(* Logix 5000 project; controller PLC_MCC1300_75F1 vendor 1 type 14 code 166 rev 32.11; software revision 32.04; part 20 of 83 *)
(* tags used below, declared in another part *)
   GP_M311A : GP_Rotator;
   M310B : MAC_Conveyor;
   M311 : MAC_Conveyor;
   M311_ALM : MAC_Conveyor_ALM;
   M311_Data : UDT_Convoy_SL;
   M311_HMR : MAC_Conveyor_HMR;
   M311_HMW : MAC_Conveyor_HMW;
   M311_M1_DR : AXIS_CIP_DRIVE;
   M311_M1_DR_IN_MAJ : MOTION_INSTRUCTION;
   M311_M1_DR_IN_MAR : MOTION_INSTRUCTION;
   M311_M1_DR_IN_MAS : MOTION_INSTRUCTION;
   M311_M1_DR_IN_MRP : MOTION_INSTRUCTION;
   M311_M1_DR_MAFR : MOTION_INSTRUCTION;
   M311_M1_DR_MDR : MOTION_INSTRUCTION;
   M311_M1_DR_MSF : MOTION_INSTRUCTION;
   M311_M1_DR_MSO : MOTION_INSTRUCTION;
   M311_M1_DR_OUT_MAJ : MOTION_INSTRUCTION;
   M311_M1_DR_OUT_MAM : MOTION_INSTRUCTION;
   M311_M1_DR_OUT_MAR : MOTION_INSTRUCTION;
   M311_M1_DR_OUT_MAS : MOTION_INSTRUCTION;
   M311_M1_DR_OUT_MCD : MOTION_INSTRUCTION;
   M311_M1_DR_OUT_MRP : MOTION_INSTRUCTION;
   M311_SpaceConv_Utilities : SpaceConv_Utilities;
   M311A : MAC_Rotator;
   M311A_HMR : MAC_Rotator_HMR;
   M311A_HMW : MAC_Rotator_HMW;
   M311A_M1_DR : AXIS_CIP_DRIVE;
   M311A_M1_DR_IN_MAM : MOTION_INSTRUCTION;
   M311A_M1_DR_IN_MAS : MOTION_INSTRUCTION;
   M311A_M1_DR_MAFR : MOTION_INSTRUCTION;
   M311A_M1_DR_MAH : MOTION_INSTRUCTION;
   M311A_M1_DR_MSF : MOTION_INSTRUCTION;
   M311A_M1_DR_MSO : MOTION_INSTRUCTION;
   M311A_M1_DR_OUT_MAJ : MOTION_INSTRUCTION;
   M311A_M1_DR_OUT_MAM : MOTION_INSTRUCTION;
   M311A_M1_DR_OUT_MAS : MOTION_INSTRUCTION;
   M311A_MAM_IP_TOFF : TIMER;
   M312 : MAC_Conveyor_Single;
   TMP_dDirection : DINT;
   TMP_r : REAL;
   TMP_rAcc : REAL;
   TMP_rDec : REAL;
   TMP_rSpeed : REAL;
   TMP_rTarget : REAL;
   TMP_rTarget_M1 : REAL;
   TMP_xForwardCommadnForCleaningZone : BOOL;
   TMP_xPositioning_M1 : BOOL;
   TMP_xPowerSaving : BOOL;
   TMP_xReverse_M1 : BOOL;
   TMP_xRun_M1 : BOOL;
   xDebugOFF : BOOL;
   Z401 : MAC_Zone;
   Z401_HMW : MAC_Zone_HMW;
(* CommandLogic, continued *)

ROUTINE M311_Output   (* ladder *)
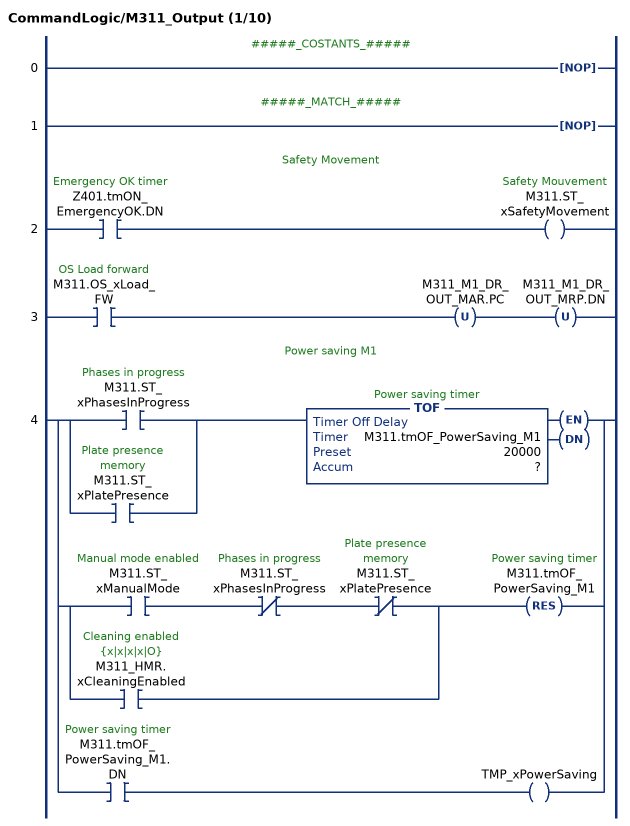
   // #####_COSTANTS_#####
   0: NOP();
   // #####_MATCH_#####
   1: NOP();
   // Safety Movement
   2: XIC(Z401.tmON_EmergencyOK.DN)OTE(M311.ST_xSafetyMovement);
   3: XIC(M311.OS_xLoad_FW)OTU(M311_M1_DR_OUT_MAR.PC)OTU(M311_M1_DR_OUT_MRP.DN);
   // Power saving M1
   4: [[XIC(M311.ST_xPhasesInProgress) ,XIC(M311.ST_xPlatePresence) ] TOF(M311.tmOF_PowerSaving_M1,?,?) ,[XIC(M311.ST_xManualMode) XIO(M311.ST_xPhasesInProgress) XIO(M311.ST_xPlatePresence) ,XIC(M311_HMR.xCleaningEnabled) ] RES(M311.tmOF_PowerSaving_M1) ,XIC(M311.tmOF_PowerSaving_M1.DN) OTE(TMP_xPowerSaving) ];
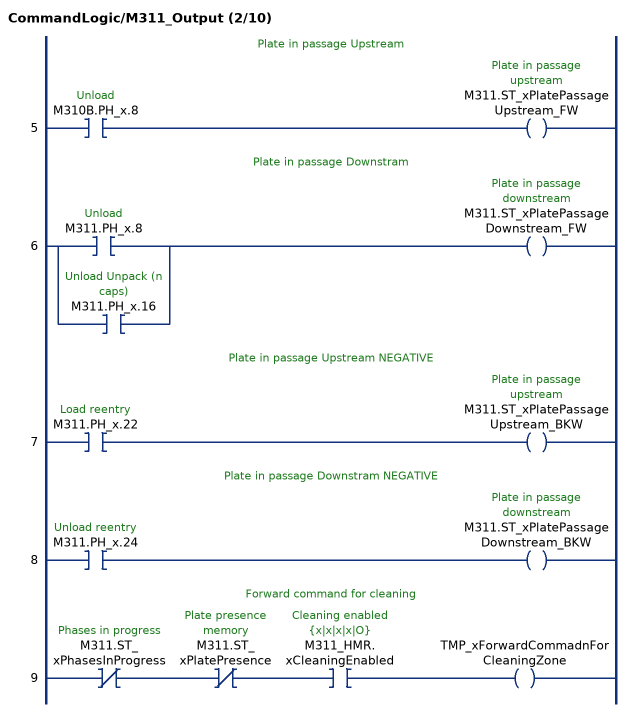
   // Plate in passage Upstream
   5: XIC(M310B.PH_x.8)OTE(M311.ST_xPlatePassageUpstream_FW);
   // Plate in passage Downstram
   6: [XIC(M311.PH_x.8) ,XIC(M311.PH_x.16) ]OTE(M311.ST_xPlatePassageDownstream_FW);
   // Plate in passage Upstream NEGATIVE
   7: XIC(M311.PH_x.22)OTE(M311.ST_xPlatePassageUpstream_BKW);
   // Plate in passage Downstram NEGATIVE
   8: XIC(M311.PH_x.24)OTE(M311.ST_xPlatePassageDownstream_BKW);
   // Forward command for cleaning
   9: XIO(M311.ST_xPhasesInProgress)XIO(M311.ST_xPlatePresence)XIC(M311_HMR.xCleaningEnabled)OTE(TMP_xForwardCommadnForCleaningZone);
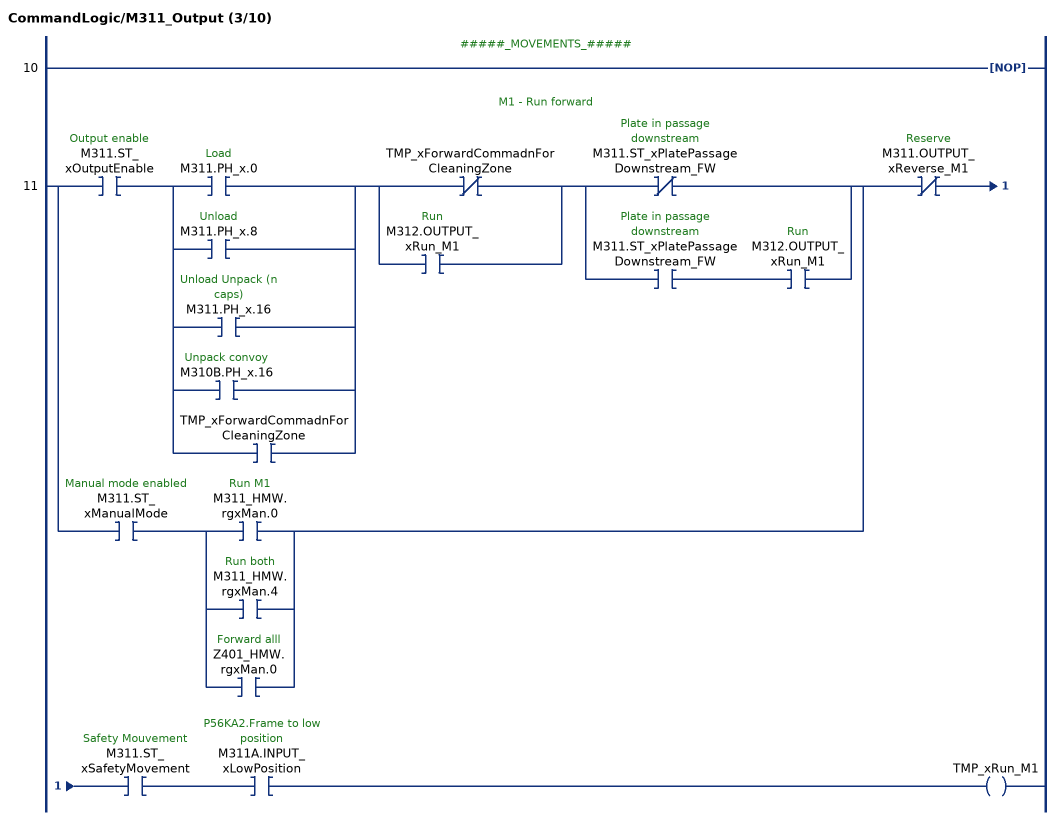
   // #####_MOVEMENTS_#####
   10: NOP();
   // M1 - Run forward
   11: [XIC(M311.ST_xOutputEnable) [XIC(M311.PH_x.0) ,XIC(M311.PH_x.8) ,XIC(M311.PH_x.16) ,XIC(M310B.PH_x.16) ,XIC(TMP_xForwardCommadnForCleaningZone) ] [XIO(TMP_xForwardCommadnForCleaningZone) ,XIC(M312.OUTPUT_xRun_M1) ] [XIO(M311.ST_xPlatePassageDownstream_FW) ,XIC(M311.ST_xPlatePassageDownstream_FW) XIC(M312.OUTPUT_xRun_M1) ] ,XIC(M311.ST_xManualMode) [XIC(M311_HMW.rgxMan.0) ,XIC(M311_HMW.rgxMan.4) ,XIC(Z401_HMW.rgxMan.0) ] ]XIO(M311.OUTPUT_xReverse_M1)XIC(M311.ST_xSafetyMovement)XIC(M311A.INPUT_xLowPosition)OTE(TMP_xRun_M1);
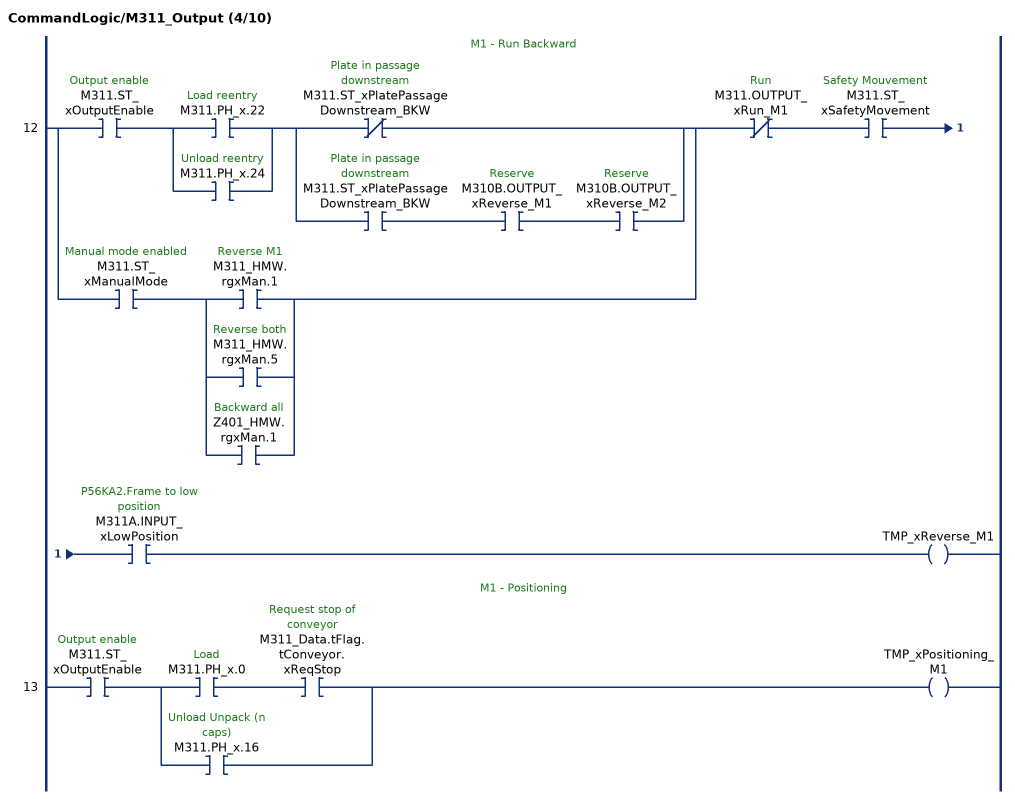
   // M1 - Run Backward
   12: [XIC(M311.ST_xOutputEnable) [XIC(M311.PH_x.22) ,XIC(M311.PH_x.24) ] [XIO(M311.ST_xPlatePassageDownstream_BKW) ,XIC(M311.ST_xPlatePassageDownstream_BKW) XIC(M310B.OUTPUT_xReverse_M1) XIC(M310B.OUTPUT_xReverse_M2) ] ,XIC(M311.ST_xManualMode) [XIC(M311_HMW.rgxMan.1) ,XIC(M311_HMW.rgxMan.5) ,XIC(Z401_HMW.rgxMan.1) ] ]XIO(M311.OUTPUT_xRun_M1)XIC(M311.ST_xSafetyMovement)XIC(M311A.INPUT_xLowPosition)OTE(TMP_xReverse_M1);
   // M1 - Positioning
   13: XIC(M311.ST_xOutputEnable)[XIC(M311.PH_x.0) XIC(M311_Data.tFlag.tConveyor.xReqStop) ,XIC(M311.PH_x.16) ]OTE(TMP_xPositioning_M1);
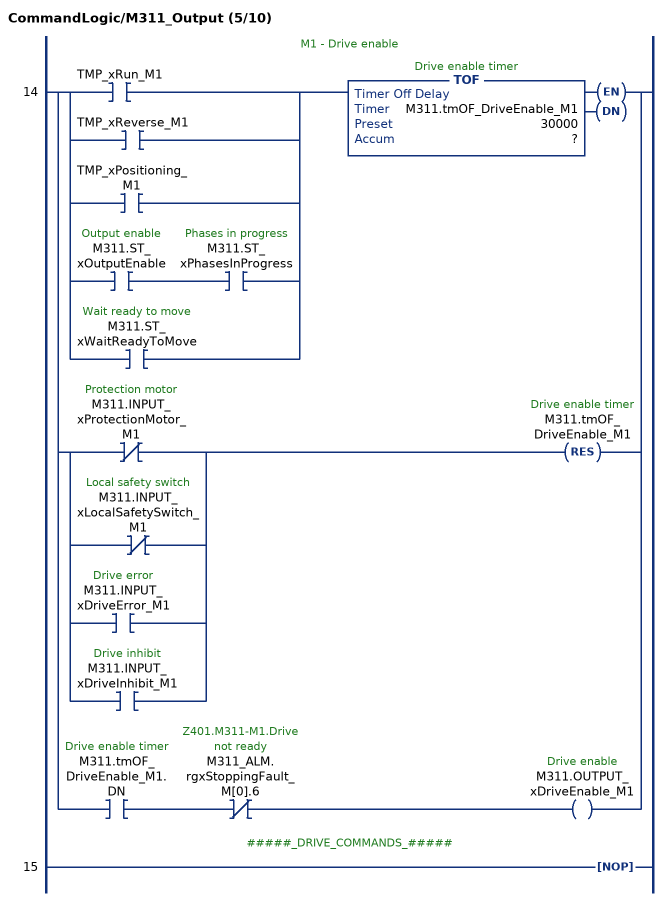
   // M1 - Drive enable
   14: [[XIC(TMP_xRun_M1) ,XIC(TMP_xReverse_M1) ,XIC(TMP_xPositioning_M1) ,XIC(M311.ST_xOutputEnable) XIC(M311.ST_xPhasesInProgress) ,XIC(M311.ST_xWaitReadyToMove) ] TOF(M311.tmOF_DriveEnable_M1,?,?) ,[XIO(M311.INPUT_xProtectionMotor_M1) ,XIO(M311.INPUT_xLocalSafetySwitch_M1) ,XIC(M311.INPUT_xDriveError_M1) ,XIC(M311.INPUT_xDriveInhibit_M1) ] RES(M311.tmOF_DriveEnable_M1) ,XIC(M311.tmOF_DriveEnable_M1.DN) XIO(M311_ALM.rgxStoppingFault_M[0].6) OTE(M311.OUTPUT_xDriveEnable_M1) ];
   // #####_DRIVE_COMMANDS_#####
   15: NOP();
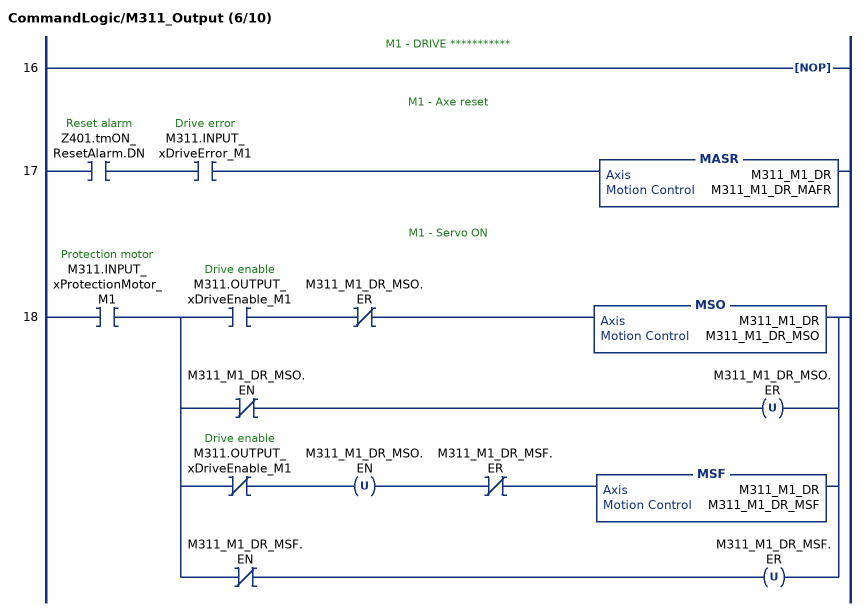
   // M1 - DRIVE ***********
   16: NOP();
   // M1 - Axe reset
   17: XIC(Z401.tmON_ResetAlarm.DN)XIC(M311.INPUT_xDriveError_M1)MASR(M311_M1_DR,M311_M1_DR_MAFR);
   // M1 - Servo ON
   18: XIC(M311.INPUT_xProtectionMotor_M1)[XIC(M311.OUTPUT_xDriveEnable_M1) XIO(M311_M1_DR_MSO.ER) MSO(M311_M1_DR,M311_M1_DR_MSO) ,XIO(M311_M1_DR_MSO.EN) OTU(M311_M1_DR_MSO.ER) ,XIO(M311.OUTPUT_xDriveEnable_M1) OTU(M311_M1_DR_MSO.EN) XIO(M311_M1_DR_MSF.ER) MSF(M311_M1_DR,M311_M1_DR_MSF) ,XIO(M311_M1_DR_MSF.EN) OTU(M311_M1_DR_MSF.ER) ];
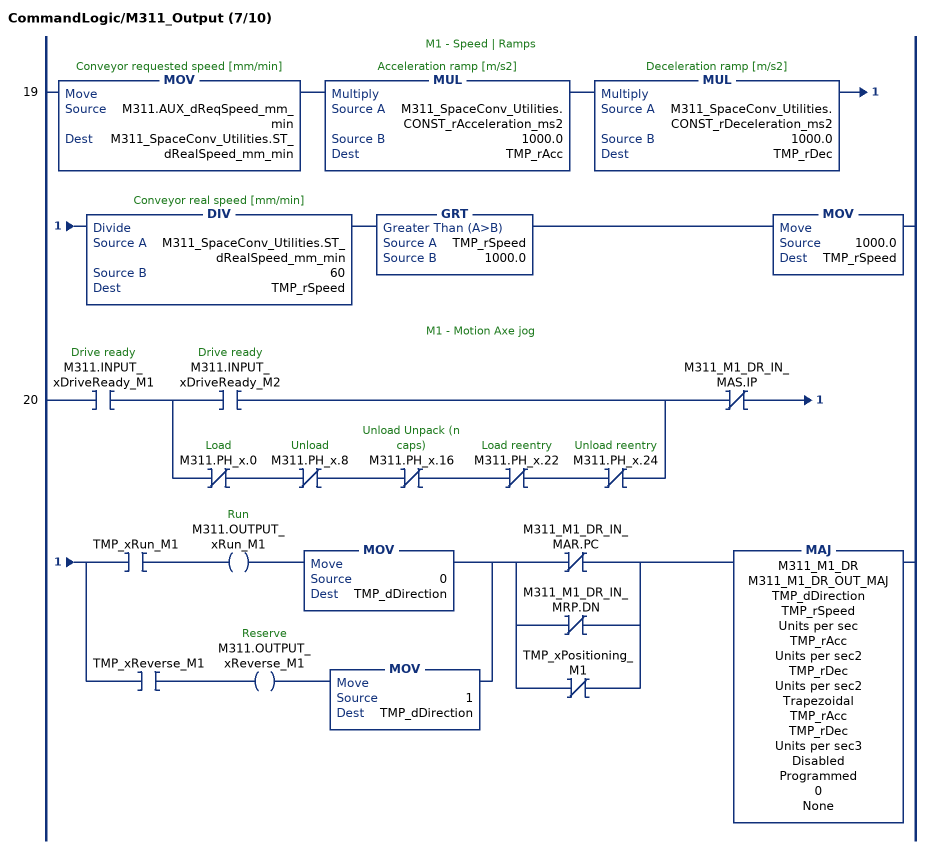
   // M1 - Speed | Ramps
   19: MOV(M311.AUX_dReqSpeed_mm_min,M311_SpaceConv_Utilities.ST_dRealSpeed_mm_min)MUL(M311_SpaceConv_Utilities.CONST_rAcceleration_ms2,1000.0,TMP_rAcc)MUL(M311_SpaceConv_Utilities.CONST_rDeceleration_ms2,1000.0,TMP_rDec)DIV(M311_SpaceConv_Utilities.ST_dRealSpeed_mm_min,60,TMP_rSpeed)GRT(TMP_rSpeed,1000.0)MOV(1000.0,TMP_rSpeed);
   // M1 - Motion Axe jog
   20: XIC(M311.INPUT_xDriveReady_M1)[XIC(M311.INPUT_xDriveReady_M2) ,XIO(M311.PH_x.0) XIO(M311.PH_x.8) XIO(M311.PH_x.16) XIO(M311.PH_x.22) XIO(M311.PH_x.24) ]XIO(M311_M1_DR_IN_MAS.IP)[XIC(TMP_xRun_M1) OTE(M311.OUTPUT_xRun_M1) MOV(0,TMP_dDirection) ,XIC(TMP_xReverse_M1) OTE(M311.OUTPUT_xReverse_M1) MOV(1,TMP_dDirection) ][XIO(M311_M1_DR_IN_MAR.PC) ,XIO(M311_M1_DR_IN_MRP.DN) ,XIO(TMP_xPositioning_M1) ]MAJ(M311_M1_DR,M311_M1_DR_OUT_MAJ,TMP_dDirection,TMP_rSpeed,Units per sec,TMP_rAcc,Units per sec2,TMP_rDec,Units per sec2,Trapezoidal,TMP_rAcc,TMP_rDec,Units per sec3,Disabled,Programmed,0,None);
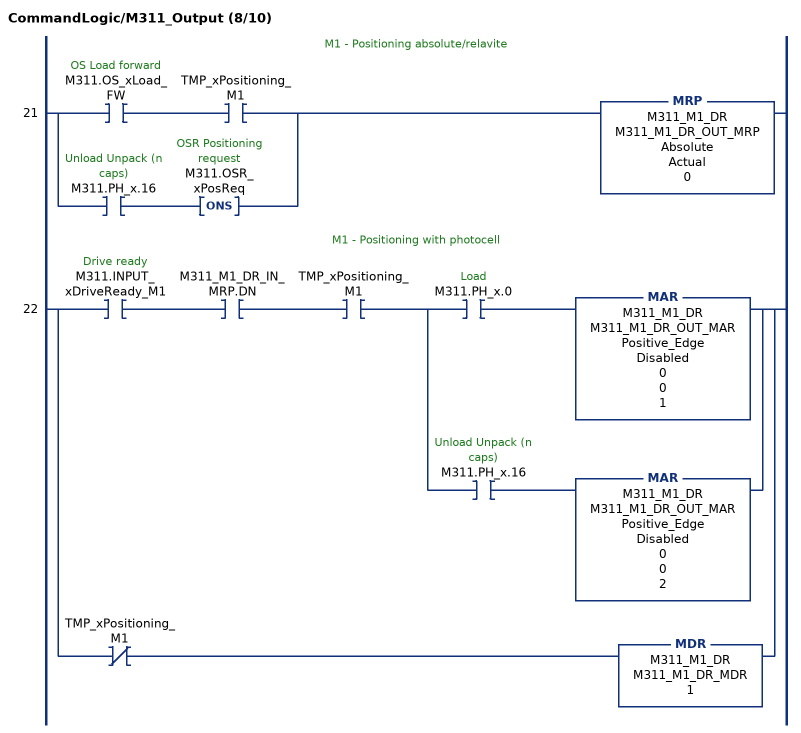
   // M1 - Positioning absolute/relavite
   21: [XIC(M311.OS_xLoad_FW) XIC(TMP_xPositioning_M1) ,XIC(M311.PH_x.16) ONS(M311.OSR_xPosReq) ]MRP(M311_M1_DR,M311_M1_DR_OUT_MRP,Absolute,Actual,0);
   // M1 - Positioning with photocell
   22: [XIC(M311.INPUT_xDriveReady_M1) XIC(M311_M1_DR_IN_MRP.DN) XIC(TMP_xPositioning_M1) [XIC(M311.PH_x.0) MAR(M311_M1_DR,M311_M1_DR_OUT_MAR,Positive_Edge,Disabled,0,0,1) ,XIC(M311.PH_x.16) MAR(M311_M1_DR,M311_M1_DR_OUT_MAR,Positive_Edge,Disabled,0,0,2) ] ,XIO(TMP_xPositioning_M1) MDR(M311_M1_DR,M311_M1_DR_MDR,1) ];
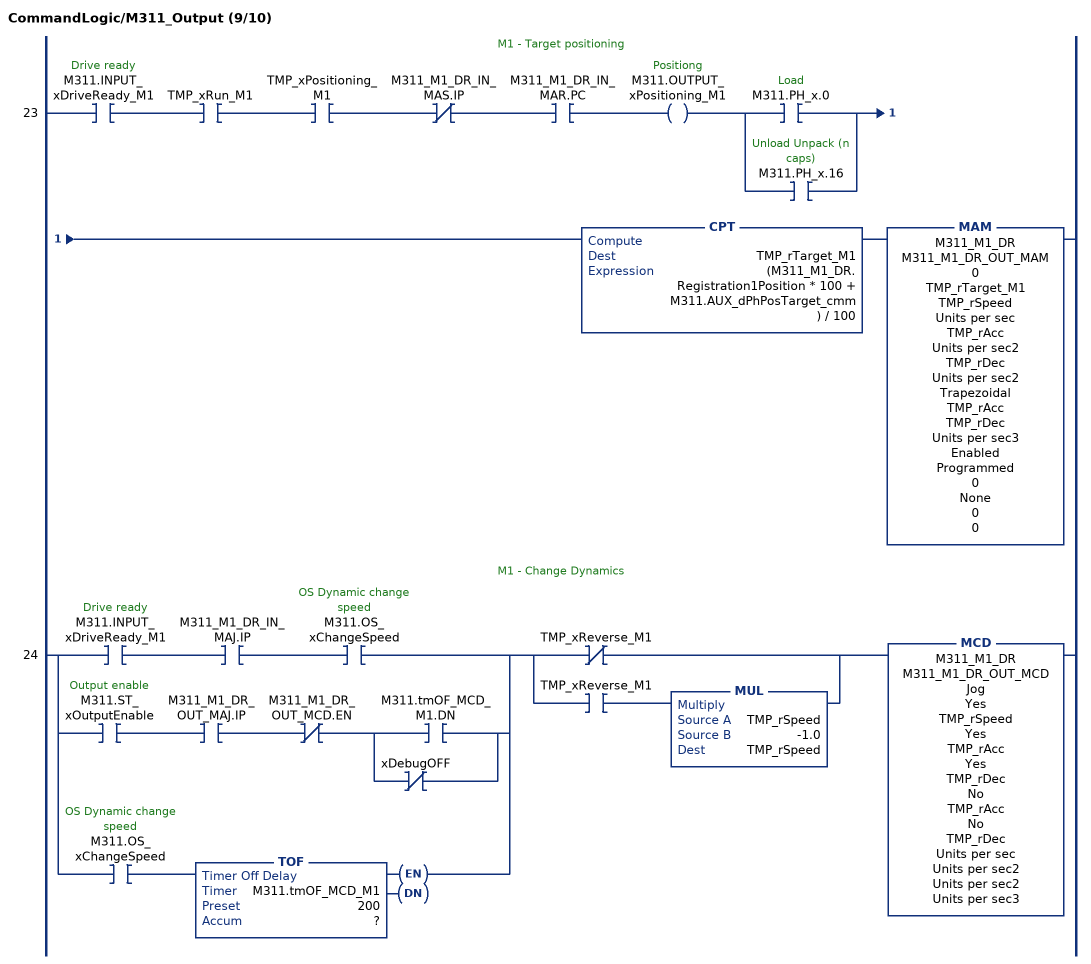
   // M1 - Target positioning
   23: XIC(M311.INPUT_xDriveReady_M1)XIC(TMP_xRun_M1)XIC(TMP_xPositioning_M1)XIO(M311_M1_DR_IN_MAS.IP)XIC(M311_M1_DR_IN_MAR.PC)OTE(M311.OUTPUT_xPositioning_M1)[XIC(M311.PH_x.0) ,XIC(M311.PH_x.16) ]CPT(TMP_rTarget_M1,(M311_M1_DR.Registration1Position * 100 + M311.AUX_dPhPosTarget_cmm ) / 100)MAM(M311_M1_DR,M311_M1_DR_OUT_MAM,0,TMP_rTarget_M1,TMP_rSpeed,Units per sec,TMP_rAcc,Units per sec2,TMP_rDec,Units per sec2,Trapezoidal,TMP_rAcc,TMP_rDec,Units per sec3,Enabled,Programmed,0,None,0,0);
   // M1 - Change Dynamics
   24: [XIC(M311.INPUT_xDriveReady_M1) XIC(M311_M1_DR_IN_MAJ.IP) XIC(M311.OS_xChangeSpeed) ,XIC(M311.ST_xOutputEnable) XIC(M311_M1_DR_OUT_MAJ.IP) XIO(M311_M1_DR_OUT_MCD.EN) [XIC(M311.tmOF_MCD_M1.DN) ,XIO(xDebugOFF) ] ,XIC(M311.OS_xChangeSpeed) TOF(M311.tmOF_MCD_M1,?,?) ][XIO(TMP_xReverse_M1) ,XIC(TMP_xReverse_M1) MUL(TMP_rSpeed,-1.0,TMP_rSpeed) ]MCD(M311_M1_DR,M311_M1_DR_OUT_MCD,Jog,Yes,TMP_rSpeed,Yes,TMP_rAcc,Yes,TMP_rDec,No,TMP_rAcc,No,TMP_rDec,Units per sec,Units per sec2,Units per sec2,Units per sec3);
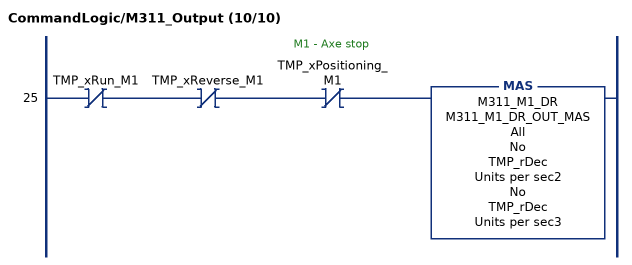
   // M1 - Axe stop
   25: XIO(TMP_xRun_M1)XIO(TMP_xReverse_M1)XIO(TMP_xPositioning_M1)MAS(M311_M1_DR,M311_M1_DR_OUT_MAS,All,No,TMP_rDec,Units per sec2,No,TMP_rDec,Units per sec3);
END_ROUTINE

ROUTINE M311A_Output   (* ladder *)
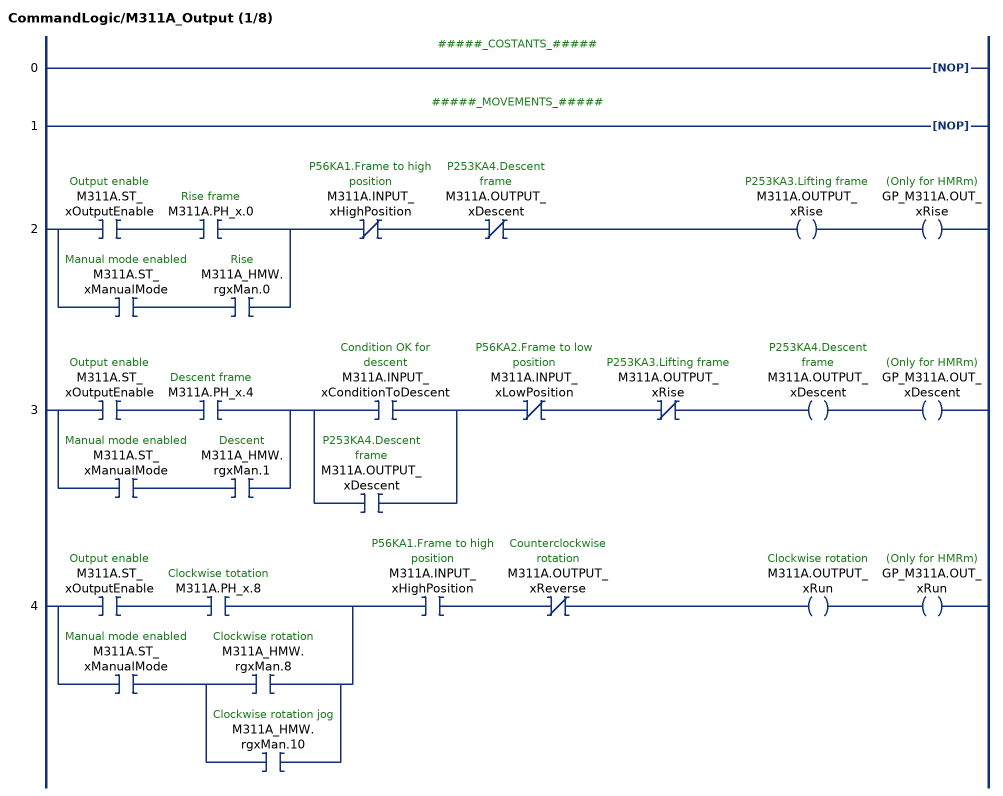
   // #####_COSTANTS_#####
   0: NOP();
   // #####_MOVEMENTS_#####
   1: NOP();
   2: [XIC(M311A.ST_xOutputEnable) XIC(M311A.PH_x.0) ,XIC(M311A.ST_xManualMode) XIC(M311A_HMW.rgxMan.0) ]XIO(M311A.INPUT_xHighPosition)XIO(M311A.OUTPUT_xDescent)OTE(M311A.OUTPUT_xRise)OTE(GP_M311A.OUT_xRise);
   3: [XIC(M311A.ST_xOutputEnable) XIC(M311A.PH_x.4) ,XIC(M311A.ST_xManualMode) XIC(M311A_HMW.rgxMan.1) ][XIC(M311A.INPUT_xConditionToDescent) ,XIC(M311A.OUTPUT_xDescent) ]XIO(M311A.INPUT_xLowPosition)XIO(M311A.OUTPUT_xRise)OTE(M311A.OUTPUT_xDescent)OTE(GP_M311A.OUT_xDescent);
   4: [XIC(M311A.ST_xOutputEnable) XIC(M311A.PH_x.8) ,XIC(M311A.ST_xManualMode) [XIC(M311A_HMW.rgxMan.8) ,XIC(M311A_HMW.rgxMan.10) ] ]XIC(M311A.INPUT_xHighPosition)XIO(M311A.OUTPUT_xReverse)OTE(M311A.OUTPUT_xRun)OTE(GP_M311A.OUT_xRun);
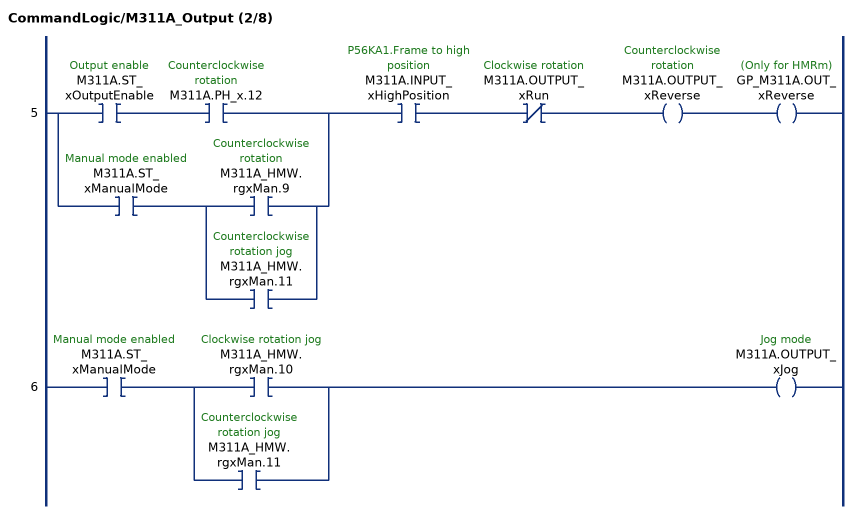
   5: [XIC(M311A.ST_xOutputEnable) XIC(M311A.PH_x.12) ,XIC(M311A.ST_xManualMode) [XIC(M311A_HMW.rgxMan.9) ,XIC(M311A_HMW.rgxMan.11) ] ]XIC(M311A.INPUT_xHighPosition)XIO(M311A.OUTPUT_xRun)OTE(M311A.OUTPUT_xReverse)OTE(GP_M311A.OUT_xReverse);
   6: XIC(M311A.ST_xManualMode)[XIC(M311A_HMW.rgxMan.10) ,XIC(M311A_HMW.rgxMan.11) ]OTE(M311A.OUTPUT_xJog);
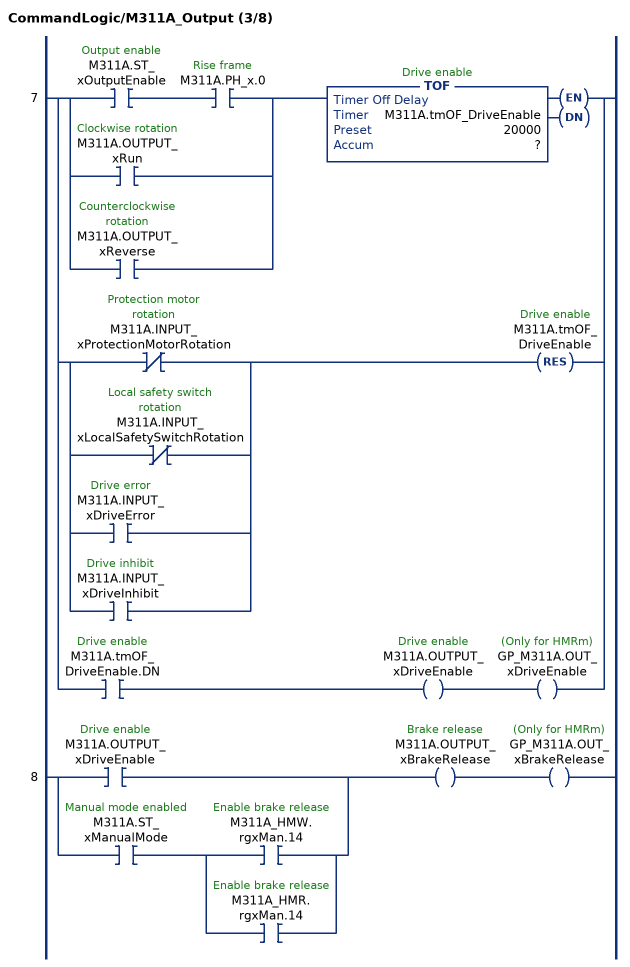
   7: [[XIC(M311A.ST_xOutputEnable) XIC(M311A.PH_x.0) ,XIC(M311A.OUTPUT_xRun) ,XIC(M311A.OUTPUT_xReverse) ] TOF(M311A.tmOF_DriveEnable,?,?) ,[XIO(M311A.INPUT_xProtectionMotorRotation) ,XIO(M311A.INPUT_xLocalSafetySwitchRotation) ,XIC(M311A.INPUT_xDriveError) ,XIC(M311A.INPUT_xDriveInhibit) ] RES(M311A.tmOF_DriveEnable) ,XIC(M311A.tmOF_DriveEnable.DN) OTE(M311A.OUTPUT_xDriveEnable) OTE(GP_M311A.OUT_xDriveEnable) ];
   8: [XIC(M311A.OUTPUT_xDriveEnable) ,XIC(M311A.ST_xManualMode) [XIC(M311A_HMW.rgxMan.14) ,XIC(M311A_HMR.rgxMan.14) ] ]OTE(M311A.OUTPUT_xBrakeRelease)OTE(GP_M311A.OUT_xBrakeRelease);
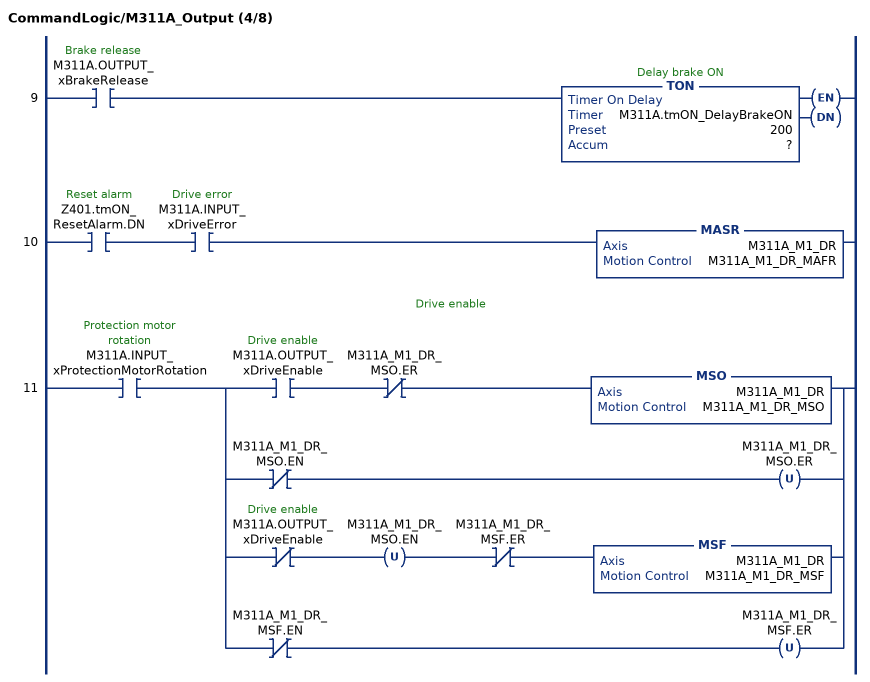
   9: XIC(M311A.OUTPUT_xBrakeRelease)TON(M311A.tmON_DelayBrakeON,?,?);
   10: XIC(Z401.tmON_ResetAlarm.DN)XIC(M311A.INPUT_xDriveError)MASR(M311A_M1_DR,M311A_M1_DR_MAFR);
   // Drive enable
   11: XIC(M311A.INPUT_xProtectionMotorRotation)[XIC(M311A.OUTPUT_xDriveEnable) XIO(M311A_M1_DR_MSO.ER) MSO(M311A_M1_DR,M311A_M1_DR_MSO) ,XIO(M311A_M1_DR_MSO.EN) OTU(M311A_M1_DR_MSO.ER) ,XIO(M311A.OUTPUT_xDriveEnable) OTU(M311A_M1_DR_MSO.EN) XIO(M311A_M1_DR_MSF.ER) MSF(M311A_M1_DR,M311A_M1_DR_MSF) ,XIO(M311A_M1_DR_MSF.EN) OTU(M311A_M1_DR_MSF.ER) ];
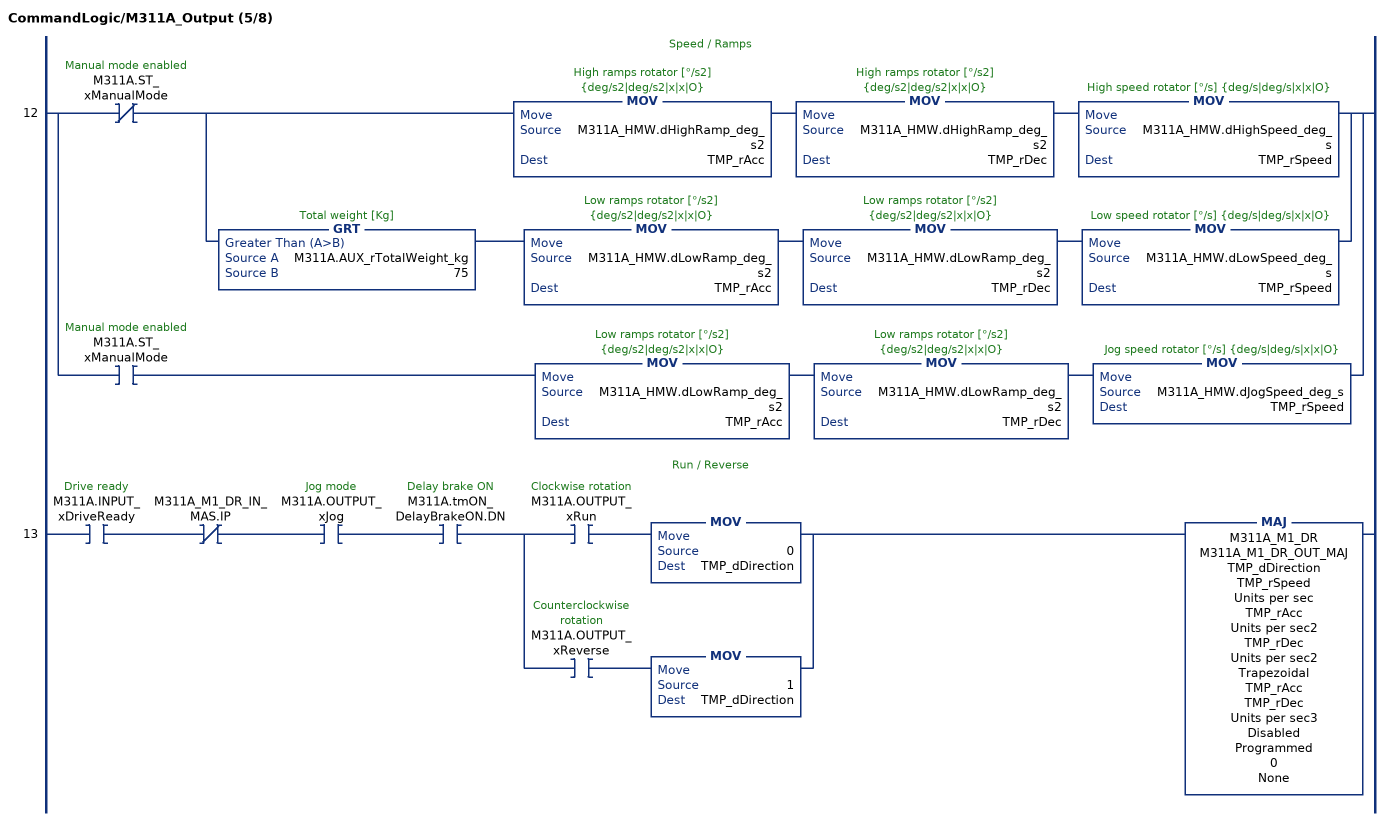
   // Speed / Ramps
   12: [XIO(M311A.ST_xManualMode) [MOV(M311A_HMW.dHighRamp_deg_s2,TMP_rAcc) MOV(M311A_HMW.dHighRamp_deg_s2,TMP_rDec) MOV(M311A_HMW.dHighSpeed_deg_s,TMP_rSpeed) ,GRT(M311A.AUX_rTotalWeight_kg,75) MOV(M311A_HMW.dLowRamp_deg_s2,TMP_rAcc) MOV(M311A_HMW.dLowRamp_deg_s2,TMP_rDec) MOV(M311A_HMW.dLowSpeed_deg_s,TMP_rSpeed) ] ,XIC(M311A.ST_xManualMode) MOV(M311A_HMW.dLowRamp_deg_s2,TMP_rAcc) MOV(M311A_HMW.dLowRamp_deg_s2,TMP_rDec) MOV(M311A_HMW.dJogSpeed_deg_s,TMP_rSpeed) ];
   // Run / Reverse
   13: XIC(M311A.INPUT_xDriveReady)XIO(M311A_M1_DR_IN_MAS.IP)XIC(M311A.OUTPUT_xJog)XIC(M311A.tmON_DelayBrakeON.DN)[XIC(M311A.OUTPUT_xRun) MOV(0,TMP_dDirection) ,XIC(M311A.OUTPUT_xReverse) MOV(1,TMP_dDirection) ]MAJ(M311A_M1_DR,M311A_M1_DR_OUT_MAJ,TMP_dDirection,TMP_rSpeed,Units per sec,TMP_rAcc,Units per sec2,TMP_rDec,Units per sec2,Trapezoidal,TMP_rAcc,TMP_rDec,Units per sec3,Disabled,Programmed,0,None);
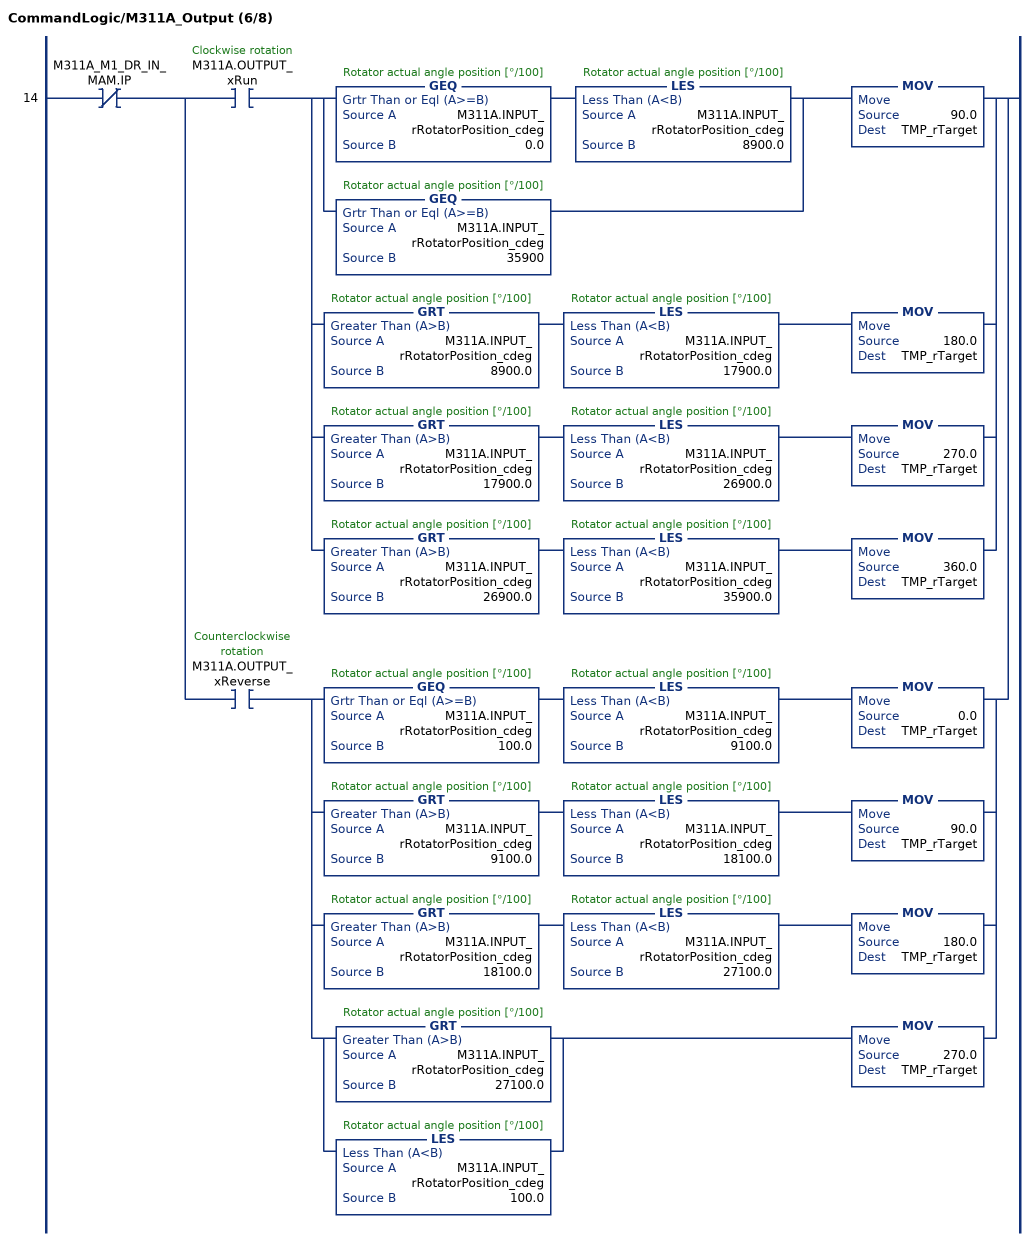
   14: XIO(M311A_M1_DR_IN_MAM.IP)[XIC(M311A.OUTPUT_xRun) [[GEQ(M311A.INPUT_rRotatorPosition_cdeg,0.0) LES(M311A.INPUT_rRotatorPosition_cdeg,8900.0) ,GEQ(M311A.INPUT_rRotatorPosition_cdeg,35900) ] MOV(90.0,TMP_rTarget) ,GRT(M311A.INPUT_rRotatorPosition_cdeg,8900.0) LES(M311A.INPUT_rRotatorPosition_cdeg,17900.0) MOV(180.0,TMP_rTarget) ,GRT(M311A.INPUT_rRotatorPosition_cdeg,17900.0) LES(M311A.INPUT_rRotatorPosition_cdeg,26900.0) MOV(270.0,TMP_rTarget) ,GRT(M311A.INPUT_rRotatorPosition_cdeg,26900.0) LES(M311A.INPUT_rRotatorPosition_cdeg,35900.0) MOV(360.0,TMP_rTarget) ] ,XIC(M311A.OUTPUT_xReverse) [GEQ(M311A.INPUT_rRotatorPosition_cdeg,100.0) LES(M311A.INPUT_rRotatorPosition_cdeg,9100.0) MOV(0.0,TMP_rTarget) ,GRT(M311A.INPUT_rRotatorPosition_cdeg,9100.0) LES(M311A.INPUT_rRotatorPosition_cdeg,18100.0) MOV(90.0,TMP_rTarget) ,GRT(M311A.INPUT_rRotatorPosition_cdeg,18100.0) LES(M311A.INPUT_rRotatorPosition_cdeg,27100.0) MOV(180.0,TMP_rTarget) ,[GRT(M311A.INPUT_rRotatorPosition_cdeg,27100.0) ,LES(M311A.INPUT_rRotatorPosition_cdeg,100.0) ] MOV(270.0,TMP_rTarget) ] ];
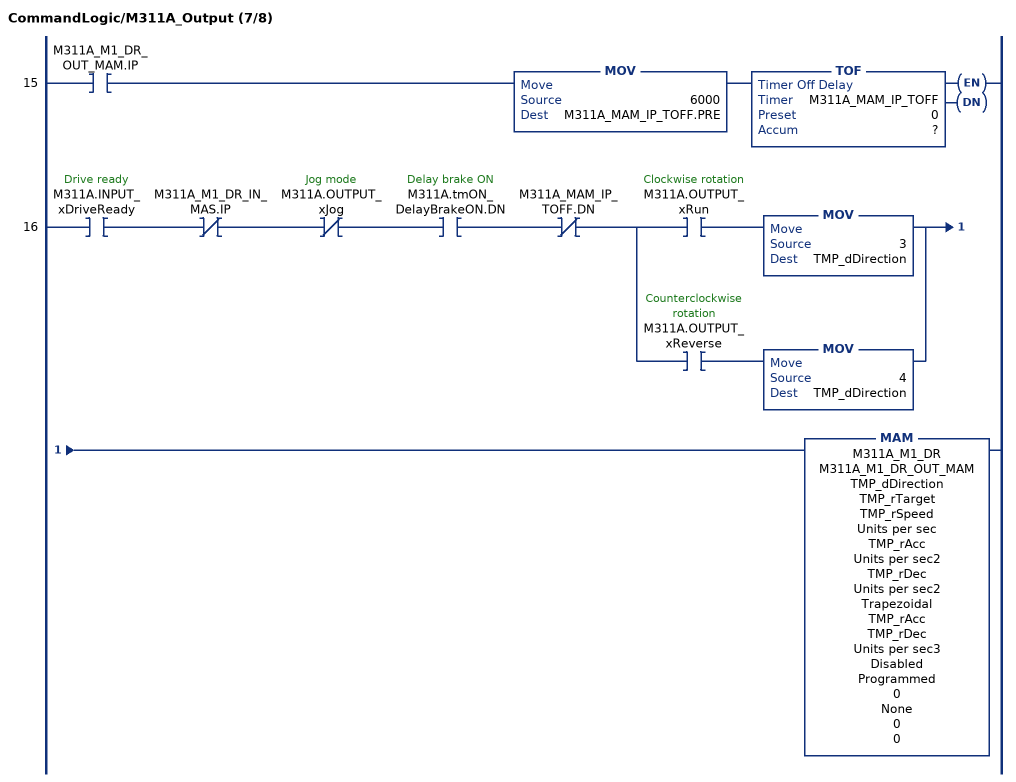
   15: XIC(M311A_M1_DR_OUT_MAM.IP)MOV(6000,M311A_MAM_IP_TOFF.PRE)TOF(M311A_MAM_IP_TOFF,?,?);
   16: XIC(M311A.INPUT_xDriveReady)XIO(M311A_M1_DR_IN_MAS.IP)XIO(M311A.OUTPUT_xJog)XIC(M311A.tmON_DelayBrakeON.DN)XIO(M311A_MAM_IP_TOFF.DN)[XIC(M311A.OUTPUT_xRun) MOV(3,TMP_dDirection) ,XIC(M311A.OUTPUT_xReverse) MOV(4,TMP_dDirection) ]MAM(M311A_M1_DR,M311A_M1_DR_OUT_MAM,TMP_dDirection,TMP_rTarget,TMP_rSpeed,Units per sec,TMP_rAcc,Units per sec2,TMP_rDec,Units per sec2,Trapezoidal,TMP_rAcc,TMP_rDec,Units per sec3,Disabled,Programmed,0,None,0,0);
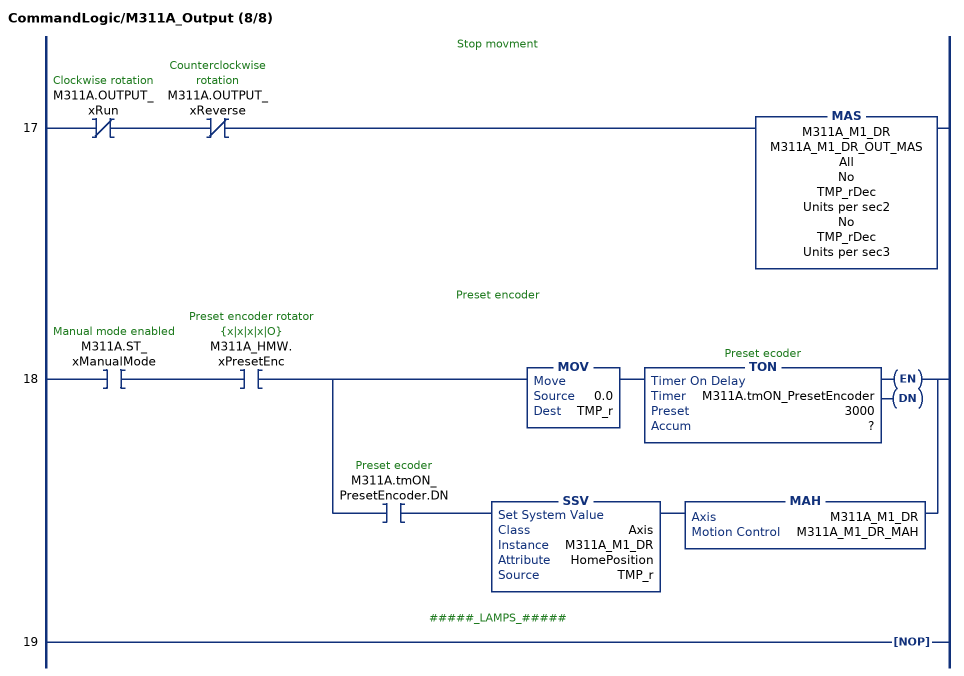
   // Stop movment
   17: XIO(M311A.OUTPUT_xRun)XIO(M311A.OUTPUT_xReverse)MAS(M311A_M1_DR,M311A_M1_DR_OUT_MAS,All,No,TMP_rDec,Units per sec2,No,TMP_rDec,Units per sec3);
   // Preset encoder
   18: XIC(M311A.ST_xManualMode)XIC(M311A_HMW.xPresetEnc)[MOV(0.0,TMP_r) TON(M311A.tmON_PresetEncoder,?,?) ,XIC(M311A.tmON_PresetEncoder.DN) SSV(Axis,M311A_M1_DR,HomePosition,TMP_r) MAH(M311A_M1_DR,M311A_M1_DR_MAH) ];
   // #####_LAMPS_#####
   19: NOP();
END_ROUTINE
